VERSION : 0.1
   VAR_INPUT
      iEnable : Bool;
      iReset : Bool;
      iAutomatic : Bool;
      iManual : Bool;
      iManualUp : Bool;
      iManualDown : Bool;
      iManualOpenForks : Bool;
      iManualCloseForks : Bool;
      iB1_up : Bool;
      iB2_mid : Bool;
      iB10 : Bool;
      iB3_dwn : Bool;
      iB5_extins : Bool;
      iB13_retras : Bool;
      iB7_palet : Bool;
      iB8_stiva : Bool;
   END_VAR
   VAR_OUTPUT
      oY4 : Bool;
      oY12 : Bool;
      oY6 : Bool;
      oY14 : Bool;
      oAlarmUpDown : Bool;
      oAlarmForks : Bool;
      oAlarmPosition : Bool;
      oAlarmFull : Bool;
   END_VAR
   VAR_IN_OUT
      xSettings : "Settings_Palletdispenser_PD2";
      xHS_PalletDispencer : "Handshakes_PalletDispenser_PD2";
   END_VAR
   VAR
      PD1 : Struct
         StepperOld : Int;
         Stepper : Int;
         MiddlePosition : Bool;
         Up : Bool;
         Down : Bool;
         Forks_In : Bool;
         Forks_Out : Bool;
      END_STRUCT;
      Alarm : Struct
         Active : Bool;
         UpDown : Bool;
         Forks : Bool;
         Position : Bool;
         Full : Bool;
      END_STRUCT;
      "Timer" : Struct
         Full : TON_TIME;
         Empty : TON_TIME;
         AlarmUpDown : TON_TIME;
         AlarmForks : TON_TIME;
      END_STRUCT;
      Flank_MiddlePosition : R_TRIG;
      Init : Bool;
   END_VAR
   VAR_TEMP
      tStep : Struct
         DISABLED : Bool;
         MANUAL : Bool;
         BLOCKED : Bool;
         IDLE : Bool;
         BASIC_POSITION : Bool;
         TO_BOTTOM_POSITION : Bool;
         FORKS_OUT_PALLET : Bool;
         WAIT_POSITION : Bool;
         TO_EMPTY_POSITION : Bool;
         EMPTY_POSITION : Bool;
         TO_MIDDLE_POSITION : Bool;
         FORKS_IN_PALLET : Bool;
         TO_UPPER_POSITION : Bool;
         FORKS_OUT_PALLET_1 : Bool;
         TO_BOTTOM_POSITION_1 : Bool;
      END_STRUCT;
   END_VAR
   VAR CONSTANT
      cSTEP_DISABLED : Int := 0;
      cSTEP_MANUAL : Int := 1;
      cSTEP_BLOCKED : Int := 7;
      cSTEP_IDLE : Int := 10;
      cSTEP_BASIC_POSITION : Int := 11;
      cSTEP_TO_MIDDLE_POSITION : Int := 12;
      cSTEP_FORKS_OUT_PALLET : Int := 13;
      cSTEP_TO_BOTTOM_POSITION : Int := 14;
      cSTEP_FORKS_IN_PALLET : Int := 15;
      cSTEP_TO_UPPER_POSITION : Int := 16;
      cSTEP_TO_BOTTOM_POSITION_1 : Int := 17;
      cSTEP_FORKS_OUT_PALLET_1 : Int := 18;
   END_VAR
BEGIN
   // ********************* INFORMATION *****************************************
   // ****************************************************************************
   // ********************* DISCLAIMER *******************************************
   // We (Qimarox) are not liable legally or in any other way for erroneous
   // program functions and their consequences!
   //    ******************** VERSION CONTROL ************************************
   //    V1.0.0 - BJA - 2018/10/22
   //    - First version of the block
   //    
   // ******************** REQUIREMENTS ******************************************
   // Data type "Handshakes_PalletDispenser_PD1"
   // Data type "Settings_Palletdispencer_PD1"
   // **************************** TO DO *****************************************
   // 
   // ****************************************************************************
   // **************************** INFO* *****************************************    
   // Pallet dispencer for picking up pallets one by one from a pallet conveyor
   // Cycle is triggered by handshaking
   // 
   // When Command.Receive is TRUE the cycle is started >> Status.Busy is TRUE
   // When cycle is completed Status.Busy is FALSE & Status.BasicPosition is TRUE
   // Pallet present must be FALSE
   // 
   // ****************************************************************************
   // ****************************************************************************
   //
   REGION Flanks
      // Positive flank middle position
      #Flank_MiddlePosition(CLK :=
                            #iB2_mid AND NOT #xSettings.Configuration.Double
                            OR
                            #iB10 AND #xSettings.Configuration.Double
      );
   END_REGION

   REGION Alarms
      REGION Alarm: Up/Down movement 
         // Reset counter if sensors are detected
         IF NOT #Alarm.UpDown THEN

            #Timer.AlarmUpDown(IN := (#iAutomatic OR #iManual) AND NOT #Alarm.UpDown AND #PD1.Up OR #PD1.Down,
                               PT := #xSettings.MaximumDurationUpDown);

            IF (#PD1.Up AND #iB1_up) OR #Flank_MiddlePosition.Q OR (#PD1.Down AND #iB3_dwn) THEN
               RESET_TIMER(#Timer.AlarmUpDown);
            END_IF;

            IF #Timer.AlarmUpDown.Q THEN
               #Alarm.UpDown := TRUE;
            END_IF;
         ELSIF #Alarm.UpDown AND #iReset THEN
            #Alarm.UpDown := FALSE;
            RESET_TIMER(#Timer.AlarmUpDown);
         END_IF;
      END_REGION
      REGION Alarm: Forks movement

         #Timer.AlarmForks(IN := (#iAutomatic OR #iManual) AND (#PD1.Forks_In OR #PD1.Forks_Out),
                           PT := #xSettings.MaximumDurationForks);


         IF NOT #Alarm.Forks THEN
            // If cilinder reaches position, reset counter
            IF (#iB5_extins AND #PD1.Forks_In OR #iB13_retras AND #PD1.Forks_Out) THEN
               RESET_TIMER(#Timer.AlarmForks);
            END_IF;
            // Create alarm if counter reaches upper time limit
            IF #Timer.AlarmForks.Q THEN
               #Alarm.Forks := TRUE;
            END_IF;

         ELSIF #Alarm.Forks AND #iReset THEN
            #Alarm.Forks := FALSE;
         END_IF;
      END_REGION
      REGION Alarm: Undefined position
         IF #Alarm.Position AND #iReset AND #iB1_up AND #iB5_extins THEN
             #Alarm.Position := FALSE;
         END_IF;
      END_REGION
      REGION Alarm: Full 
         #Timer.Full(IN := #iB8_stiva AND NOT #Alarm.Full,
                     PT := T#2S);
         #Timer.Empty(IN := NOT #iB8_stiva AND #Alarm.Full,
                      PT := T#5s);

         IF NOT #Alarm.Full AND #iB1_up AND #Timer.Full.Q THEN
            #Alarm.Full := TRUE;
         ELSIF #Alarm.Full AND #Timer.Empty.Q THEN
            #Alarm.Full := FALSE;
         END_IF;
      END_REGION
      REGION Alarm: Active
         #Alarm.Active :=
         #Alarm.UpDown OR
         #Alarm.Forks OR
         #Alarm.Position
         ;
      END_REGION
   END_REGION
   REGION Make active steps bits
      // This ensures only one step is possible every cpu cycle
      #tStep.DISABLED := #PD1.Stepper = #cSTEP_DISABLED;
      #tStep.MANUAL := #PD1.Stepper = #cSTEP_MANUAL;
      #tStep.BLOCKED := #PD1.Stepper = #cSTEP_BLOCKED;
      #tStep.IDLE := #PD1.Stepper = #cSTEP_IDLE;
      #tStep.BASIC_POSITION := #PD1.Stepper = #cSTEP_BASIC_POSITION;
      #tStep.TO_MIDDLE_POSITION := #PD1.Stepper = #cSTEP_TO_MIDDLE_POSITION;
      #tStep.FORKS_OUT_PALLET := #PD1.Stepper = #cSTEP_FORKS_OUT_PALLET;
      #tStep.TO_BOTTOM_POSITION := #PD1.Stepper = #cSTEP_TO_BOTTOM_POSITION;
      #tStep.FORKS_IN_PALLET := #PD1.Stepper = #cSTEP_FORKS_IN_PALLET;
      #tStep.TO_UPPER_POSITION := #PD1.Stepper = #cSTEP_TO_UPPER_POSITION;
      #tStep.FORKS_OUT_PALLET_1 := #PD1.Stepper = #cSTEP_FORKS_OUT_PALLET_1;
      #tStep.TO_BOTTOM_POSITION_1 := #PD1.Stepper = #cSTEP_TO_BOTTOM_POSITION_1;
   END_REGION
   REGION Step 0: Disabled
      IF #PD1.Stepper = #cSTEP_DISABLED THEN
         IF #tStep.DISABLED THEN

            // Handshake signals
            #xHS_PalletDispencer.Status.Blocked := TRUE;
            #xHS_PalletDispencer.Status.Busy := FALSE;
            #xHS_PalletDispencer.Status.BasicPosition := FALSE;
            #xHS_PalletDispencer.Status.WaitPosition := FALSE;

            // Movements
            #PD1.Up := FALSE;
            #PD1.Down := FALSE;
            #PD1.Forks_In := FALSE;
            #PD1.Forks_Out := FALSE;

            // Module enabled 
            IF #iEnable THEN
               // Installation is in manual mode
               // go to manual step
               IF #iManual THEN
                  #PD1.Stepper := #cSTEP_MANUAL;
               // Installation is in automatic mode
               // go to idle step
               ELSIF #iAutomatic THEN
                  #PD1.Stepper := #cSTEP_IDLE;
               END_IF;
            END_IF;
         END_IF;
      ELSE
         IF NOT #iEnable THEN
            #PD1.Stepper := #cSTEP_DISABLED;
         END_IF;
      END_IF;
   END_REGION
   REGION Step 1: Manual
       IF #Alarm.Active AND #PD1.Stepper <> #cSTEP_MANUAL THEN
           #PD1.StepperOld := #PD1.Stepper;
           #PD1.Stepper := #cSTEP_MANUAL;
       END_IF;
      IF #PD1.Stepper = #cSTEP_MANUAL THEN
         IF #tStep.MANUAL THEN

            // Handshake signals
            #xHS_PalletDispencer.Status.Blocked := TRUE;
            #xHS_PalletDispencer.Status.Busy := FALSE;
            #xHS_PalletDispencer.Status.BasicPosition := FALSE;
            #xHS_PalletDispencer.Status.WaitPosition := FALSE;

            REGION Stop at middle position
               IF (#iManualUp OR #iManualDown) AND #Flank_MiddlePosition.Q AND NOT #PD1.MiddlePosition THEN
                  #PD1.MiddlePosition := TRUE;
               ELSIF NOT #iManualUp AND NOT #iManualDown AND #PD1.MiddlePosition THEN
                  #PD1.MiddlePosition := FALSE;
               END_IF;
            END_REGION
            REGION Movement up
               #PD1.Up := #iManualUp AND NOT #iManualDown AND NOT #iB1_up AND NOT #PD1.MiddlePosition;
            END_REGION
            REGION Movement down
               #PD1.Down := #iManualDown AND NOT #iManualUp AND NOT #iB3_dwn AND NOT #PD1.MiddlePosition;
            END_REGION
            REGION Forks in pallet
               #PD1.Forks_In := #iManualCloseForks AND NOT #iB5_extins;
            END_REGION
            REGION Forks out pallet
               #PD1.Forks_Out := #iManualOpenForks AND NOT #iB13_retras;
            END_REGION
            REGION Manual disabled
                IF NOT #iManual AND NOT #Alarm.Active THEN //zz
                  #PD1.Stepper := #cSTEP_DISABLED;
               END_IF;
            END_REGION
         END_IF;
      END_IF;
   END_REGION
   REGION Step 7: Blocked
     /// IF #Alarm.Active AND #PD1.Stepper <> #cSTEP_BLOCKED THEN
      //   #PD1.StepperOld := #PD1.Stepper;
     //    #PD1.Stepper := #cSTEP_BLOCKED;
     // END_IF;

      IF #PD1.Stepper = #cSTEP_BLOCKED THEN
          IF #tStep.BLOCKED THEN

              // Handshake signals
              #xHS_PalletDispencer.Status.Blocked := TRUE;
              #xHS_PalletDispencer.Status.Busy := FALSE;
              #xHS_PalletDispencer.Status.BasicPosition := FALSE;
              #xHS_PalletDispencer.Status.WaitPosition := FALSE;

              // Movements
              #PD1.Up := FALSE;
              #PD1.Down := FALSE;
              #PD1.Forks_In := FALSE;
              #PD1.Forks_Out := FALSE;
              IF #iManual THEN
                  #PD1.Forks_In := #iManualCloseForks AND NOT #iB5_extins;//zz
                  #PD1.Up := #iManualUp AND NOT #iManualDown AND NOT (#iB1_up OR #iB2_mid);// zz
              END_IF;
              IF #Init THEN
                  #PD1.Forks_In := #Init AND NOT #iB5_extins;
                  #PD1.Up := #Init AND #iB5_extins AND NOT #iB1_up;// zz
              END_IF;

              // Alarms resolved
              IF NOT #Alarm.Active THEN
                  #PD1.Stepper := #cSTEP_DISABLED;
              END_IF;
          END_IF;
      END_IF;
   END_REGION
   REGION Step 10: Idle
      IF #PD1.Stepper = #cSTEP_IDLE THEN
         IF #tStep.IDLE THEN

            // Handshake signals
            #xHS_PalletDispencer.Status.Blocked := FALSE;
            #xHS_PalletDispencer.Status.Busy := FALSE;
            #xHS_PalletDispencer.Status.BasicPosition := FALSE;
            #xHS_PalletDispencer.Status.WaitPosition := FALSE;

            // Movements
            #PD1.Up := FALSE;
            #PD1.Down := FALSE;
            #PD1.Forks_In := FALSE;
            #PD1.Forks_Out := FALSE;

            // Check position
            // 
            // Basic position; 
            // Upper position & forks in palletstack
            IF #iB1_up AND #iB5_extins THEN
               #PD1.Stepper := #cSTEP_BASIC_POSITION;
            // Middle position
            ELSIF (
               #iB2_mid AND NOT #xSettings.Configuration.Double
               OR
               #iB10 AND #xSettings.Configuration.Double
               )
            THEN
               // Forks in pallet stack
               IF #iB5_extins THEN
                  IF #iB7_palet THEN
                     #PD1.Stepper := #cSTEP_FORKS_OUT_PALLET;
                  ELSE
                     #PD1.Stepper := #cSTEP_TO_UPPER_POSITION;
                  END_IF;
               // Forks out pallet stack
               ELSIF #iB13_retras THEN
                  #PD1.Stepper := #cSTEP_TO_BOTTOM_POSITION;
               ELSE
                  #Alarm.Position := TRUE;
               END_IF;
            // Bottom position
            ELSIF #iB3_dwn THEN
               // Forks in pallet stack
               IF #iB5_extins THEN
                  #PD1.Stepper := #cSTEP_TO_UPPER_POSITION;
               // Forks out pallet stack
               ELSIF #iB13_retras THEN
                  #PD1.Stepper := #cSTEP_FORKS_IN_PALLET;
               ELSE
                  #Alarm.Position := TRUE;
               END_IF;
            // If forks are in palletstack and not at upper/middle/bottom position, then go back to basic position 
            ELSIF #iB5_extins THEN
               #PD1.Stepper := #cSTEP_TO_UPPER_POSITION;
            ELSE
               #Alarm.Position := TRUE;
            END_IF;

            IF NOT #iAutomatic THEN
               #PD1.StepperOld := #PD1.Stepper;
               #PD1.Stepper := #cSTEP_DISABLED;
            END_IF;
         END_IF;
      END_IF;
   END_REGION
   REGION Step 11: Basic position
      IF #PD1.Stepper = #cSTEP_BASIC_POSITION THEN
         IF #tStep.BASIC_POSITION THEN

            // Handshake signals
            #xHS_PalletDispencer.Status.Blocked := FALSE;
            #xHS_PalletDispencer.Status.Busy := FALSE;
            #xHS_PalletDispencer.Status.BasicPosition := TRUE;
            #xHS_PalletDispencer.Status.WaitPosition := FALSE;

            // Movements
            #PD1.Up := FALSE;
            #PD1.Down := FALSE;
            #PD1.Forks_In := FALSE;
            #PD1.Forks_Out := FALSE;


            // Basic position; 
            // Upper position & forks in palletstack
            IF #iAutomatic THEN
               // If command receive is high 
               IF #xHS_PalletDispencer.Command.Receive
                  // Requested pallettype must match with configured pallettype
                  AND #xHS_PalletDispencer.Command.Pallettype = #xSettings.Configuration.Pallettype
                  // and pallet is detected
                  AND #iB7_palet
               THEN
                  #PD1.Stepper := #cSTEP_TO_MIDDLE_POSITION;
              END_IF;
              IF #xHS_PalletDispencer.Command.Deliver THEN
                  #PD1.Stepper := #cSTEP_TO_BOTTOM_POSITION_1;
              END_IF;
            END_IF;

            IF NOT #iAutomatic THEN
               #PD1.StepperOld := #PD1.Stepper;
               #PD1.Stepper := #cSTEP_DISABLED;
            END_IF;
         END_IF;
      END_IF;
   END_REGION
   REGION Step 12: Move to middle position
      IF #PD1.Stepper = #cSTEP_TO_MIDDLE_POSITION THEN
         IF #tStep.TO_MIDDLE_POSITION THEN

            // Handshake signals
            #xHS_PalletDispencer.Status.Blocked := FALSE;
            #xHS_PalletDispencer.Status.Busy := TRUE;
            #xHS_PalletDispencer.Status.BasicPosition := FALSE;
            #xHS_PalletDispencer.Status.WaitPosition := FALSE;

            // Movements
            #PD1.Up := FALSE;
            #PD1.Down := TRUE;
            #PD1.Forks_In := FALSE;
            #PD1.Forks_Out := FALSE;

            // If command is given to pickup pallet stack 
            // go to forks in pallet
            IF #iB2_mid AND NOT #xSettings.Configuration.Double THEN
               #PD1.Stepper := #cSTEP_FORKS_OUT_PALLET;
            ELSIF #iB10 AND #xSettings.Configuration.Double THEN
               #PD1.Stepper := #cSTEP_FORKS_OUT_PALLET;
            END_IF;

            IF NOT #iAutomatic THEN
               #PD1.StepperOld := #PD1.Stepper;
               #PD1.Stepper := #cSTEP_DISABLED;
            END_IF;
         END_IF;
      END_IF;
   END_REGION
   REGION Step 13: Move forks out of pallet
      IF #PD1.Stepper = #cSTEP_FORKS_OUT_PALLET THEN
         IF #tStep.FORKS_OUT_PALLET THEN

            // Handshake signals
            #xHS_PalletDispencer.Status.Blocked := FALSE;
            #xHS_PalletDispencer.Status.Busy := TRUE;
            #xHS_PalletDispencer.Status.BasicPosition := FALSE;
            #xHS_PalletDispencer.Status.WaitPosition := FALSE;

            // Movements
            #PD1.Up := FALSE;
            #PD1.Down := FALSE;
            #PD1.Forks_In := FALSE;
            #PD1.Forks_Out := TRUE;

            // If forks are out of palletstack
            // then wait position is reached
            IF #iB13_retras THEN
               #PD1.Stepper := #cSTEP_TO_BOTTOM_POSITION;
            END_IF;

            IF NOT #iAutomatic THEN
               #PD1.StepperOld := #PD1.Stepper;
               #PD1.Stepper := #cSTEP_DISABLED;
            END_IF;
         END_IF;
      END_IF;
   END_REGION
   REGION Step 14: Movement to bottom position
      IF #PD1.Stepper = #cSTEP_TO_BOTTOM_POSITION THEN
         IF #tStep.TO_BOTTOM_POSITION THEN

            // Handshake signals
            #xHS_PalletDispencer.Status.Blocked := FALSE;
            #xHS_PalletDispencer.Status.Busy := TRUE;
            #xHS_PalletDispencer.Status.BasicPosition := FALSE;
            #xHS_PalletDispencer.Status.WaitPosition := FALSE;

            // Movements
            #PD1.Up := FALSE;
            #PD1.Down := TRUE;
            #PD1.Forks_In := FALSE;
            #PD1.Forks_Out := FALSE;

            // If bottom position is reached, then move out forks
            IF #iB3_dwn THEN
               #PD1.Stepper := #cSTEP_FORKS_IN_PALLET;
            END_IF;

            IF NOT #iAutomatic THEN
               #PD1.StepperOld := #PD1.Stepper;
               #PD1.Stepper := #cSTEP_DISABLED;
            END_IF;
         END_IF;
      END_IF;
   END_REGION
   REGION Step 15: Move forks in pallet
      IF #PD1.Stepper = #cSTEP_FORKS_IN_PALLET THEN
         IF #tStep.FORKS_IN_PALLET THEN

            // Handshake signals
            #xHS_PalletDispencer.Status.Blocked := FALSE;
            #xHS_PalletDispencer.Status.Busy := TRUE;
            #xHS_PalletDispencer.Status.BasicPosition := FALSE;
            #xHS_PalletDispencer.Status.WaitPosition := FALSE;

            // Movements
            #PD1.Up := FALSE;
            #PD1.Down := FALSE;
            #PD1.Forks_In := TRUE;
            #PD1.Forks_Out := FALSE;

            // If forks are in pallet stack
            // go to upper position
            IF #iB5_extins THEN
               #PD1.Stepper := #cSTEP_TO_UPPER_POSITION;
            END_IF;

            IF NOT #iAutomatic THEN
               #PD1.StepperOld := #PD1.Stepper;
               #PD1.Stepper := #cSTEP_DISABLED;
            END_IF;
         END_IF;
      END_IF;
   END_REGION
   REGION Step 16: Move to upper position
      IF #PD1.Stepper = #cSTEP_TO_UPPER_POSITION THEN
         IF #tStep.TO_UPPER_POSITION THEN

            // Handshake signals
            #xHS_PalletDispencer.Status.Blocked := FALSE;
            #xHS_PalletDispencer.Status.Busy := TRUE;
            #xHS_PalletDispencer.Status.BasicPosition := FALSE;
            #xHS_PalletDispencer.Status.WaitPosition := FALSE;

            // Movements
            #PD1.Up := TRUE;
            #PD1.Down := FALSE;
            #PD1.Forks_In := FALSE;
            #PD1.Forks_Out := FALSE;

            // If in upper position
            IF #iB1_up THEN
               #PD1.Stepper := #cSTEP_IDLE;
            END_IF;

            IF NOT #iAutomatic THEN
               #PD1.StepperOld := #PD1.Stepper;
               #PD1.Stepper := #cSTEP_DISABLED;
            END_IF;
         END_IF;
      END_IF;
   END_REGION
   REGION Step 17: Move to bottom-delivery
       IF #PD1.Stepper = #cSTEP_TO_BOTTOM_POSITION_1   THEN
           IF #tStep.TO_BOTTOM_POSITION_1 THEN

               // Handshake signals
               #xHS_PalletDispencer.Status.Blocked := FALSE;
               #xHS_PalletDispencer.Status.Busy := TRUE;
               #xHS_PalletDispencer.Status.BasicPosition := FALSE;
               #xHS_PalletDispencer.Status.WaitPosition := FALSE;

               // Movements
               #PD1.Up := false;
               #PD1.Down := true;
               #PD1.Forks_In := FALSE;
               #PD1.Forks_Out := FALSE;

               // If in upper position
                   IF #iB3_dwn THEN
                       #PD1.Stepper := #cSTEP_FORKS_OUT_PALLET_1;

               END_IF;

               IF NOT #iAutomatic THEN
                   #PD1.StepperOld := #PD1.Stepper;
                   #PD1.Stepper := #cSTEP_DISABLED;
               END_IF;
           END_IF;
       END_IF;
   END_REGION
   REGION Step 18: Fork out-delivery
       IF #PD1.Stepper = #cSTEP_FORKS_OUT_PALLET_1 THEN
           IF #tStep.FORKS_OUT_PALLET_1 THEN

               // Handshake signals
               #xHS_PalletDispencer.Status.Blocked := FALSE;
               #xHS_PalletDispencer.Status.Busy := TRUE;
               #xHS_PalletDispencer.Status.BasicPosition := FALSE;
               #xHS_PalletDispencer.Status.WaitPosition := FALSE;

               // Movements
               #PD1.Up := false;
               #PD1.Down := false;
               #PD1.Forks_In := FALSE;
               #PD1.Forks_Out := true;

               // If in upper position
               IF #iB13_retras AND NOT  #xHS_PalletDispencer.Command.Deliver THEN 
             //      #PD1.Stepper := #cSTEP_IDLE;
                  ;
               END_IF;

               IF NOT #iAutomatic THEN
                   #PD1.StepperOld := #PD1.Stepper;
                   #PD1.Stepper := #cSTEP_DISABLED;
               END_IF;
           END_IF;
       END_IF;
   END_REGION
   REGION Movements
      // Movements
      #oY4 := #PD1.Up;
      #oY12 := #PD1.Down;
      #oY6 := #PD1.Forks_In;
      #oY14 := #PD1.Forks_Out;
   END_REGION
   REGION Alarm feedback
      #oAlarmUpDown := #Alarm.UpDown;
      #oAlarmForks := #Alarm.Forks;
      #oAlarmPosition := #Alarm.Position;
      #oAlarmFull := #Alarm.Full;
   END_REGION
   REGION Status handshakes
      #xHS_PalletDispencer.Status.PalletPresent := #iB7_palet AND #xHS_PalletDispencer.Status.BasicPosition;
      #xHS_PalletDispencer.Status.Pallettype := #xSettings.Configuration.Pallettype;
      #xHS_PalletDispencer.Status.Step := #PD1.Stepper;
   END_REGION
END_FUNCTION_BLOCK

FUNCTION "FC_AckOpTranzit" : Void   // FC1, SCL
{ S7_Optimized_Access := 'TRUE' }
VERSION : 0.1
   VAR_TEMP
      i : Int;
      almw : Word;
   END_VAR
BEGIN
   "HMI".tip_sel := 0;
   "HMI".instance_sel := 0;
   "HMI".msop_vizi := 0;
   FOR #i := 0 TO 6 DO
       #almw := "s".f[#i].almw;
       IF (#almw<> 0) THEN
           IF #almw.%X3 THEN
               "HMI".tip_sel := 1;
               "HMI".msop_vizi := 1;
           END_IF;
           IF #almw.%X2 THEN
               "HMI".tip_sel := 2;
               "HMI".msop_vizi := 2;
           END_IF;
           IF (#almw.%X0 OR #almw.%X1 ) THEN
               "HMI".tip_sel := 3;
               "HMI".msop_vizi := 3;
           END_IF;
           "HMI".instance_sel := #i;
       END_IF;
   END_FOR;


   "HMI".chg_prio := false;
   IF "HMI".tip_sel <> "HMI".tip_sel_v OR "HMI".instance_sel <> "HMI".instance_sel_v THEN
       "HMI".tip_sel_v := "HMI".tip_sel;
       "HMI".instance_sel_v := "HMI".instance_sel;
       "HMI".chg_prio := TRUE;
       "HMI".ButOpMem := 0;
   END_IF;
   "HMI".ButOpW := 0;
   IF "HMI".ButOpHMI <> 0 THEN
       "HMI".ButOpW := "HMI".ButOpHMI;
       "HMI".ButOpHMI := 0;
       "HMI".ButOpMem := "HMI".ButOpW;
   END_IF;

   "HMI".ButOpVis := 7;
   "HMI".numSt := "HMI".instance_sel;
END_FUNCTION

FUNCTION "FC60_MappingIn" : Void   // FC2, LAD
{ S7_Optimized_Access := 'TRUE' }
VERSION : 0.1
   VAR_TEMP
      pulse_bit : Bool;
   END_VAR
   VAR_TEMP   // added for the SCL form of the ladder/FBD networks
      _w1 : Bool;
   END_VAR
BEGIN

REGION Network 1
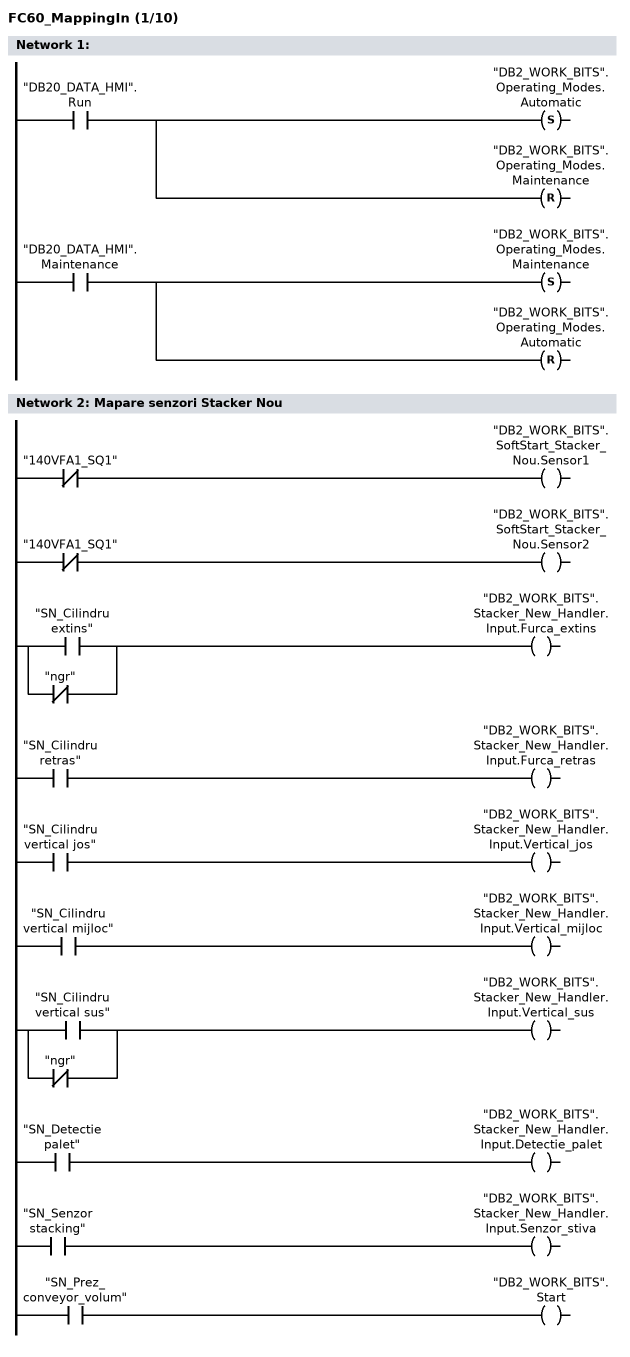
   RUNG wire#powerrail
      Contact( "DB20_DATA_HMI".Run )
      wire#w1
      S_Coil( "DB2_WORK_BITS".Operating_Modes.Automatic )
   END_RUNG
   RUNG wire#w1
      R_Coil( "DB2_WORK_BITS".Operating_Modes.Maintenance )
   END_RUNG
   RUNG wire#powerrail
      Contact( "DB20_DATA_HMI".Maintenance )
      wire#w2
      S_Coil( "DB2_WORK_BITS".Operating_Modes.Maintenance )
   END_RUNG
   RUNG wire#w2
      R_Coil( "DB2_WORK_BITS".Operating_Modes.Automatic )
   END_RUNG
   // the same network as SCL:
   IF "DB20_DATA_HMI".Run THEN
       "DB2_WORK_BITS".Operating_Modes.Automatic := TRUE;
       "DB2_WORK_BITS".Operating_Modes.Maintenance := FALSE;
   END_IF;
   IF "DB20_DATA_HMI".Maintenance THEN
       "DB2_WORK_BITS".Operating_Modes.Maintenance := TRUE;
       "DB2_WORK_BITS".Operating_Modes.Automatic := FALSE;
   END_IF;
END_REGION

REGION Network 2: Mapare senzori Stacker Nou
   RUNG wire#powerrail
      I_Contact( "140VFA1_SQ1" )
      Coil( "DB2_WORK_BITS".SoftStart_Stacker_Nou.Sensor1 )
   END_RUNG
   RUNG wire#powerrail
      I_Contact( "140VFA1_SQ1" )
      Coil( "DB2_WORK_BITS".SoftStart_Stacker_Nou.Sensor2 )
   END_RUNG
   RUNG wire#powerrail
      Contact( "SN_Cilindru extins" )
      wire#w1
      Coil( "DB2_WORK_BITS".Stacker_New_Handler.Input.Furca_extins )
   END_RUNG
   RUNG wire#powerrail
      I_Contact( "ngr" )
   END_RUNG wire#w1
   RUNG wire#powerrail
      Contact( "SN_Cilindru retras" )
      Coil( "DB2_WORK_BITS".Stacker_New_Handler.Input.Furca_retras )
   END_RUNG
   RUNG wire#powerrail
      Contact( "SN_Cilindru vertical jos" )
      Coil( "DB2_WORK_BITS".Stacker_New_Handler.Input.Vertical_jos )
   END_RUNG
   RUNG wire#powerrail
      Contact( "SN_Cilindru vertical mijloc" )
      Coil( "DB2_WORK_BITS".Stacker_New_Handler.Input.Vertical_mijloc )
   END_RUNG
   RUNG wire#powerrail
      Contact( "SN_Cilindru vertical sus" )
      wire#w2
      Coil( "DB2_WORK_BITS".Stacker_New_Handler.Input.Vertical_sus )
   END_RUNG
   RUNG wire#powerrail
      I_Contact( "ngr" )
   END_RUNG wire#w2
   RUNG wire#powerrail
      Contact( "SN_Detectie palet" )
      Coil( "DB2_WORK_BITS".Stacker_New_Handler.Input.Detectie_palet )
   END_RUNG
   RUNG wire#powerrail
      Contact( "SN_Senzor stacking" )
      Coil( "DB2_WORK_BITS".Stacker_New_Handler.Input.Senzor_stiva )
   END_RUNG
   RUNG wire#powerrail
      Contact( "SN_Prez_conveyor_volum" )
      Coil( "DB2_WORK_BITS".Start )
   END_RUNG
   // the same network as SCL:
   "DB2_WORK_BITS".SoftStart_Stacker_Nou.Sensor1 := NOT "140VFA1_SQ1";
   "DB2_WORK_BITS".SoftStart_Stacker_Nou.Sensor2 := NOT "140VFA1_SQ1";
   "DB2_WORK_BITS".Stacker_New_Handler.Input.Furca_extins := "SN_Cilindru extins" OR NOT "ngr";
   "DB2_WORK_BITS".Stacker_New_Handler.Input.Furca_retras := "SN_Cilindru retras";
   "DB2_WORK_BITS".Stacker_New_Handler.Input.Vertical_jos := "SN_Cilindru vertical jos";
   "DB2_WORK_BITS".Stacker_New_Handler.Input.Vertical_mijloc := "SN_Cilindru vertical mijloc";
   "DB2_WORK_BITS".Stacker_New_Handler.Input.Vertical_sus := "SN_Cilindru vertical sus" OR NOT "ngr";
   "DB2_WORK_BITS".Stacker_New_Handler.Input.Detectie_palet := "SN_Detectie palet";
   "DB2_WORK_BITS".Stacker_New_Handler.Input.Senzor_stiva := "SN_Senzor stacking";
   "DB2_WORK_BITS".Start := "SN_Prez_conveyor_volum";
END_REGION

REGION Network 3: Mapare senzori Stacker Nou
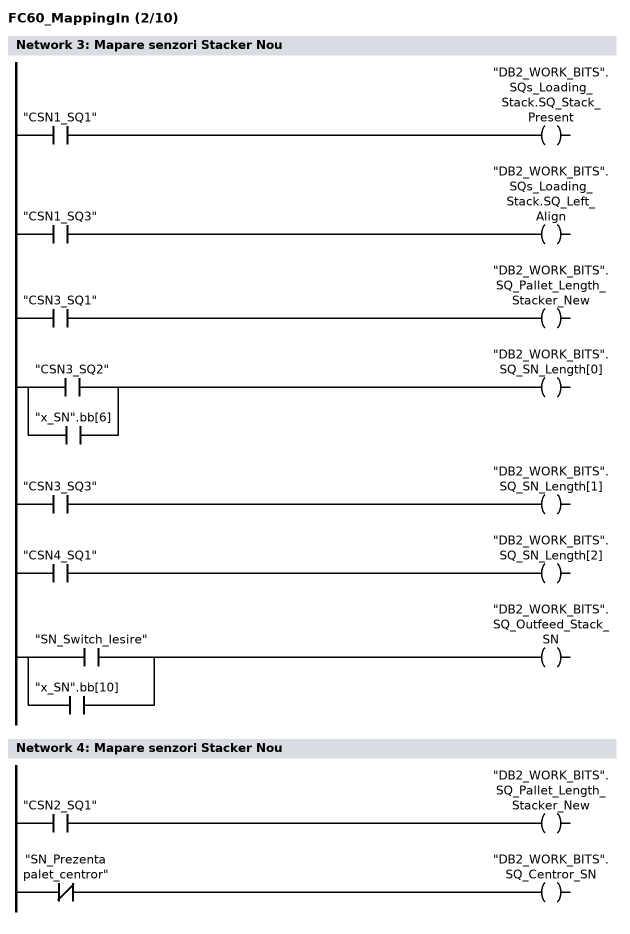
   RUNG wire#powerrail
      Contact( "CSN1_SQ1" )
      Coil( "DB2_WORK_BITS".SQs_Loading_Stack.SQ_Stack_Present )
   END_RUNG
   RUNG wire#powerrail
      Contact( "CSN1_SQ3" )
      Coil( "DB2_WORK_BITS".SQs_Loading_Stack.SQ_Left_Align )
   END_RUNG
   RUNG wire#powerrail
      Contact( "CSN3_SQ1" )
      Coil( "DB2_WORK_BITS".SQ_Pallet_Length_Stacker_New )
   END_RUNG
   RUNG wire#powerrail
      Contact( "CSN3_SQ2" )
      wire#w1
      Coil( "DB2_WORK_BITS".SQ_SN_Length[0] )
   END_RUNG
   RUNG wire#powerrail
      Contact( "x_SN".bb[6] )
   END_RUNG wire#w1
   RUNG wire#powerrail
      Contact( "CSN3_SQ3" )
      Coil( "DB2_WORK_BITS".SQ_SN_Length[1] )
   END_RUNG
   RUNG wire#powerrail
      Contact( "CSN4_SQ1" )
      Coil( "DB2_WORK_BITS".SQ_SN_Length[2] )
   END_RUNG
   RUNG wire#powerrail
      Contact( "SN_Switch_Iesire" )
      wire#w2
      Coil( "DB2_WORK_BITS".SQ_Outfeed_Stack_SN )
   END_RUNG
   RUNG wire#powerrail
      Contact( "x_SN".bb[10] )
   END_RUNG wire#w2
   // the same network as SCL:
   "DB2_WORK_BITS".SQs_Loading_Stack.SQ_Stack_Present := "CSN1_SQ1";
   "DB2_WORK_BITS".SQs_Loading_Stack.SQ_Left_Align := "CSN1_SQ3";
   "DB2_WORK_BITS".SQ_Pallet_Length_Stacker_New := "CSN3_SQ1";
   "DB2_WORK_BITS".SQ_SN_Length[0] := "CSN3_SQ2" OR "x_SN".bb[6];
   "DB2_WORK_BITS".SQ_SN_Length[1] := "CSN3_SQ3";
   "DB2_WORK_BITS".SQ_SN_Length[2] := "CSN4_SQ1";
   "DB2_WORK_BITS".SQ_Outfeed_Stack_SN := "SN_Switch_Iesire" OR "x_SN".bb[10];
END_REGION

REGION Network 4: Mapare senzori Stacker Nou
   RUNG wire#powerrail
      Contact( "CSN2_SQ1" )
      Coil( "DB2_WORK_BITS".SQ_Pallet_Length_Stacker_New )
   END_RUNG
   RUNG wire#powerrail
      I_Contact( "SN_Prezenta palet_centror" )
      Coil( "DB2_WORK_BITS".SQ_Centror_SN )
   END_RUNG
   // the same network as SCL:
   "DB2_WORK_BITS".SQ_Pallet_Length_Stacker_New := "CSN2_SQ1";
   "DB2_WORK_BITS".SQ_Centror_SN := NOT "SN_Prezenta palet_centror";
END_REGION

REGION Network 5: Mapare senzori Stacker
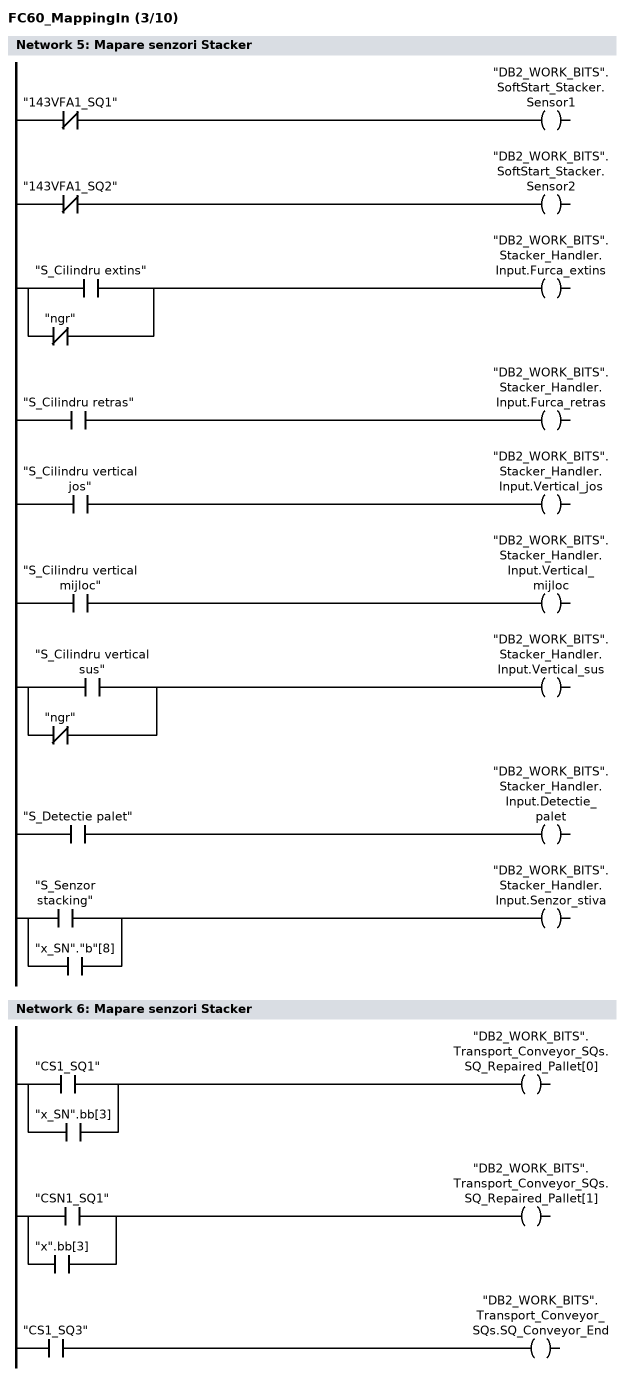
   RUNG wire#powerrail
      I_Contact( "143VFA1_SQ1" )
      Coil( "DB2_WORK_BITS".SoftStart_Stacker.Sensor1 )
   END_RUNG
   RUNG wire#powerrail
      I_Contact( "143VFA1_SQ2" )
      Coil( "DB2_WORK_BITS".SoftStart_Stacker.Sensor2 )
   END_RUNG
   RUNG wire#powerrail
      Contact( "S_Cilindru extins" )
      wire#w1
      Coil( "DB2_WORK_BITS".Stacker_Handler.Input.Furca_extins )
   END_RUNG
   RUNG wire#powerrail
      I_Contact( "ngr" )
   END_RUNG wire#w1
   RUNG wire#powerrail
      Contact( "S_Cilindru retras" )
      Coil( "DB2_WORK_BITS".Stacker_Handler.Input.Furca_retras )
   END_RUNG
   RUNG wire#powerrail
      Contact( "S_Cilindru vertical jos" )
      Coil( "DB2_WORK_BITS".Stacker_Handler.Input.Vertical_jos )
   END_RUNG
   RUNG wire#powerrail
      Contact( "S_Cilindru vertical mijloc" )
      Coil( "DB2_WORK_BITS".Stacker_Handler.Input.Vertical_mijloc )
   END_RUNG
   RUNG wire#powerrail
      Contact( "S_Cilindru vertical sus" )
      wire#w2
      Coil( "DB2_WORK_BITS".Stacker_Handler.Input.Vertical_sus )
   END_RUNG
   RUNG wire#powerrail
      I_Contact( "ngr" )
   END_RUNG wire#w2
   RUNG wire#powerrail
      Contact( "S_Detectie palet" )
      Coil( "DB2_WORK_BITS".Stacker_Handler.Input.Detectie_palet )
   END_RUNG
   RUNG wire#powerrail
      Contact( "S_Senzor stacking" )
      wire#w3
      Coil( "DB2_WORK_BITS".Stacker_Handler.Input.Senzor_stiva )
   END_RUNG
   RUNG wire#powerrail
      Contact( "x_SN"."b"[8] )
   END_RUNG wire#w3
   // the same network as SCL:
   "DB2_WORK_BITS".SoftStart_Stacker.Sensor1 := NOT "143VFA1_SQ1";
   "DB2_WORK_BITS".SoftStart_Stacker.Sensor2 := NOT "143VFA1_SQ2";
   "DB2_WORK_BITS".Stacker_Handler.Input.Furca_extins := "S_Cilindru extins" OR NOT "ngr";
   "DB2_WORK_BITS".Stacker_Handler.Input.Furca_retras := "S_Cilindru retras";
   "DB2_WORK_BITS".Stacker_Handler.Input.Vertical_jos := "S_Cilindru vertical jos";
   "DB2_WORK_BITS".Stacker_Handler.Input.Vertical_mijloc := "S_Cilindru vertical mijloc";
   "DB2_WORK_BITS".Stacker_Handler.Input.Vertical_sus := "S_Cilindru vertical sus" OR NOT "ngr";
   "DB2_WORK_BITS".Stacker_Handler.Input.Detectie_palet := "S_Detectie palet";
   "DB2_WORK_BITS".Stacker_Handler.Input.Senzor_stiva := "S_Senzor stacking" OR "x_SN"."b"[8];
END_REGION

REGION Network 6: Mapare senzori Stacker
   RUNG wire#powerrail
      Contact( "CS1_SQ1" )
      wire#w1
      Coil( "DB2_WORK_BITS".Transport_Conveyor_SQs.SQ_Repaired_Pallet[0] )
   END_RUNG
   RUNG wire#powerrail
      Contact( "x_SN".bb[3] )
   END_RUNG wire#w1
   RUNG wire#powerrail
      Contact( "CSN1_SQ1" )
      wire#w2
      Coil( "DB2_WORK_BITS".Transport_Conveyor_SQs.SQ_Repaired_Pallet[1] )
   END_RUNG
   RUNG wire#powerrail
      Contact( "x".bb[3] )
   END_RUNG wire#w2
   RUNG wire#powerrail
      Contact( "CS1_SQ3" )
      Coil( "DB2_WORK_BITS".Transport_Conveyor_SQs.SQ_Conveyor_End )
   END_RUNG
   // the same network as SCL:
   "DB2_WORK_BITS".Transport_Conveyor_SQs.SQ_Repaired_Pallet[0] := "CS1_SQ1" OR "x_SN".bb[3];
   "DB2_WORK_BITS".Transport_Conveyor_SQs.SQ_Repaired_Pallet[1] := "CSN1_SQ1" OR "x".bb[3];
   "DB2_WORK_BITS".Transport_Conveyor_SQs.SQ_Conveyor_End := "CS1_SQ3";
END_REGION

REGION Network 7: Mapare senzori Stacker
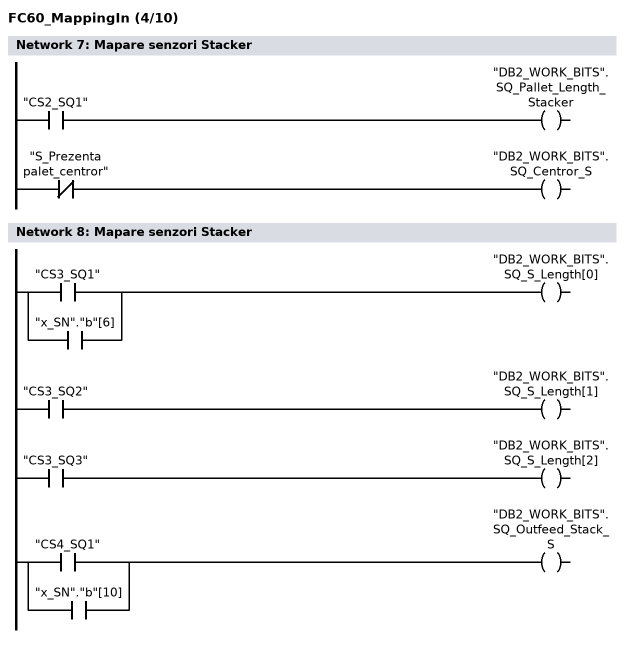
   RUNG wire#powerrail
      Contact( "CS2_SQ1" )
      Coil( "DB2_WORK_BITS".SQ_Pallet_Length_Stacker )
   END_RUNG
   RUNG wire#powerrail
      I_Contact( "S_Prezenta palet_centror" )
      Coil( "DB2_WORK_BITS".SQ_Centror_S )
   END_RUNG
   // the same network as SCL:
   "DB2_WORK_BITS".SQ_Pallet_Length_Stacker := "CS2_SQ1";
   "DB2_WORK_BITS".SQ_Centror_S := NOT "S_Prezenta palet_centror";
END_REGION

REGION Network 8: Mapare senzori Stacker
   RUNG wire#powerrail
      Contact( "CS3_SQ1" )
      wire#w1
      Coil( "DB2_WORK_BITS".SQ_S_Length[0] )
   END_RUNG
   RUNG wire#powerrail
      Contact( "x_SN"."b"[6] )
   END_RUNG wire#w1
   RUNG wire#powerrail
      Contact( "CS3_SQ2" )
      Coil( "DB2_WORK_BITS".SQ_S_Length[1] )
   END_RUNG
   RUNG wire#powerrail
      Contact( "CS3_SQ3" )
      Coil( "DB2_WORK_BITS".SQ_S_Length[2] )
   END_RUNG
   RUNG wire#powerrail
      Contact( "CS4_SQ1" )
      wire#w2
      Coil( "DB2_WORK_BITS".SQ_Outfeed_Stack_S )
   END_RUNG
   RUNG wire#powerrail
      Contact( "x_SN"."b"[10] )
   END_RUNG wire#w2
   // the same network as SCL:
   "DB2_WORK_BITS".SQ_S_Length[0] := "CS3_SQ1" OR "x_SN"."b"[6];
   "DB2_WORK_BITS".SQ_S_Length[1] := "CS3_SQ2";
   "DB2_WORK_BITS".SQ_S_Length[2] := "CS3_SQ3";
   "DB2_WORK_BITS".SQ_Outfeed_Stack_S := "CS4_SQ1" OR "x_SN"."b"[10];
END_REGION

